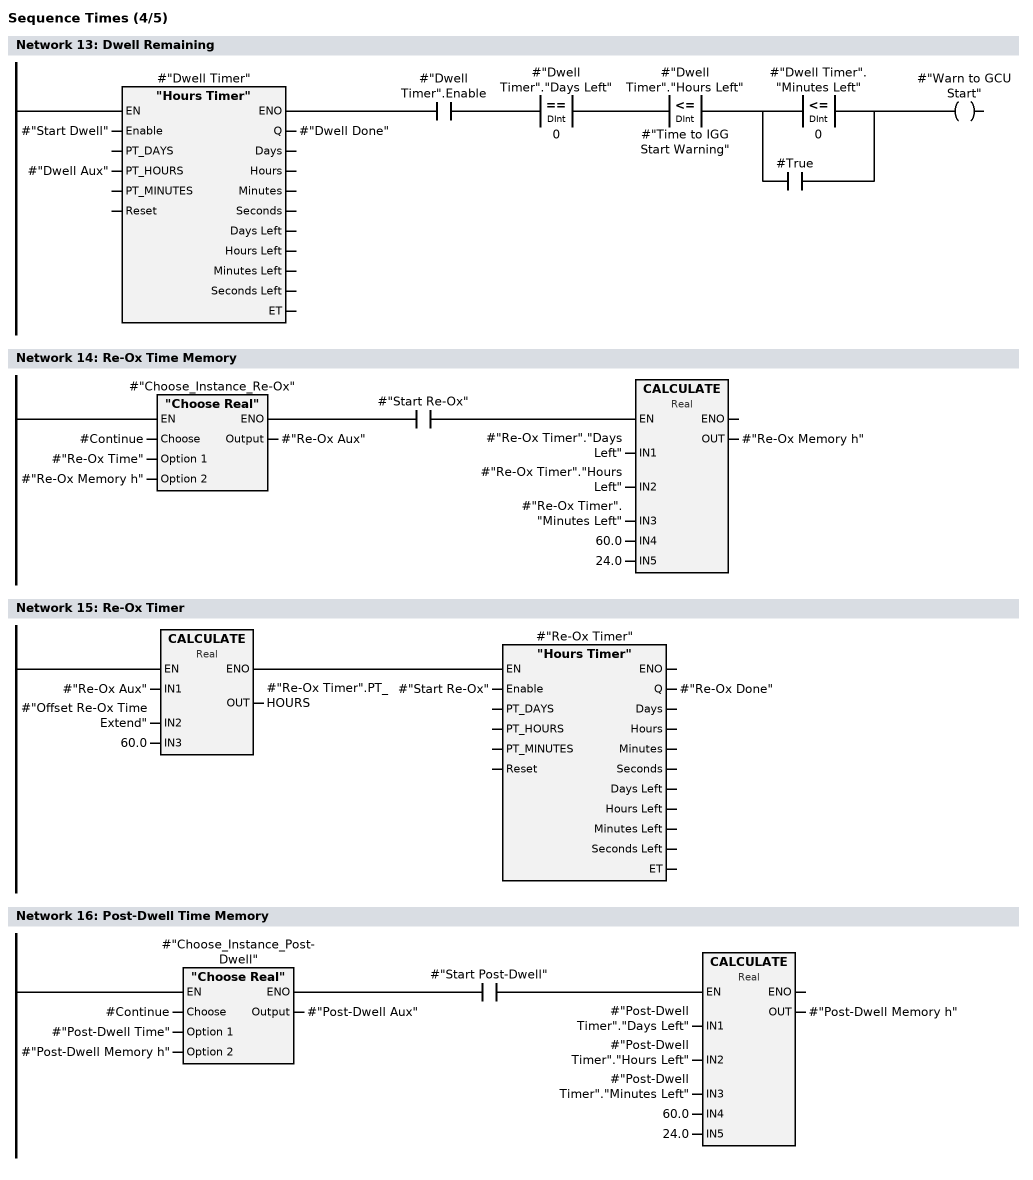
   RUNG wire#powerrail
      #"Dwell Timer"(Enable := #"Start Dwell", PT_DAYS :=, PT_HOURS := #"Dwell Aux", PT_MINUTES :=, Reset :=, Q => #"Dwell Done", Days =>, Hours =>, Minutes =>, Seconds =>, "Days Left" =>, "Hours Left" =>, "Minutes Left" =>, "Seconds Left" =>, ET =>)
      Contact( #"Dwell Timer".Enable )
      { S7_Templates := "SrcType := DInt" } EQ_Contact(in1 := #"Dwell Timer"."Days Left", in2 := 0)
      { S7_Templates := "SrcType := DInt" } LE_Contact(in1 := #"Dwell Timer"."Hours Left", in2 := #"Time to IGG Start Warning")
      wire#w1
      { S7_Templates := "SrcType := DInt" } LE_Contact(in1 := #"Dwell Timer"."Minutes Left", in2 := 0)
      wire#w2
      Coil( #"Warn to GCU Start" )
   END_RUNG
   RUNG wire#w1
      Contact( #True )
   END_RUNG wire#w2
   // the same network as SCL:
   #"Dwell Timer"(Enable := #"Start Dwell", PT_HOURS := #"Dwell Aux", Q => #"Dwell Done", ENO => #_w1);   // "Hours Timer"
   #"Warn to GCU Start" := #_w1 AND #"Dwell Timer".Enable AND (#"Dwell Timer"."Days Left" = 0) AND (#"Dwell Timer"."Hours Left" <= #"Time to IGG Start Warning") AND ((#"Dwell Timer"."Minutes Left" <= 0) OR #True);
END_REGION

REGION Network 14: Re-Ox Time Memory
   RUNG wire#powerrail
      #"Choose_Instance_Re-Ox"(Choose := #Continue, "Option 1" := #"Re-Ox Time", "Option 2" := #"Re-Ox Memory h", Output => #"Re-Ox Aux")
      Contact( #"Start Re-Ox" )
      { S7_Templates := "SrcType := Real"; S7_Expression := "(IN1*IN5)+IN2+(IN3/IN4)" } Calculate(in1 := #"Re-Ox Timer"."Days Left", in2 := #"Re-Ox Timer"."Hours Left", in3 := #"Re-Ox Timer"."Minutes Left", in4 := 60.0, in5 := 24.0, out => #"Re-Ox Memory h")
   END_RUNG
   // the same network as SCL:
   #"Choose_Instance_Re-Ox"(Choose := #Continue,   // "Choose Real"
                           "Option 1" := #"Re-Ox Time",
                           "Option 2" := #"Re-Ox Memory h",
                           Output => #"Re-Ox Aux",
                           ENO => #_w1);
   IF #_w1 AND #"Start Re-Ox" THEN
       #"Re-Ox Memory h" := (#"Re-Ox Timer"."Days Left"*24.0)+#"Re-Ox Timer"."Hours Left"+(#"Re-Ox Timer"."Minutes Left"/60.0);
   END_IF;
END_REGION

REGION Network 15: Re-Ox Timer
   RUNG wire#powerrail
      { S7_Templates := "SrcType := Real"; S7_Expression := "IN1+IN2" } Calculate(in1 := #"Re-Ox Aux", in2 := #"Offset Re-Ox Time Extend", in3 := 60.0, out => #"Re-Ox Timer".PT_HOURS)
      #"Re-Ox Timer"(Enable := #"Start Re-Ox", PT_DAYS :=, PT_HOURS :=, PT_MINUTES :=, Reset :=, Q => #"Re-Ox Done", Days =>, Hours =>, Minutes =>, Seconds =>, "Days Left" =>, "Hours Left" =>, "Minutes Left" =>, "Seconds Left" =>, ET =>)
   END_RUNG
   // the same network as SCL:
   #"Re-Ox Timer".PT_HOURS := #"Re-Ox Aux"+#"Offset Re-Ox Time Extend";
   #"Re-Ox Timer"(Enable := #"Start Re-Ox", Q => #"Re-Ox Done");   // "Hours Timer"
END_REGION

REGION Network 16: Post-Dwell Time Memory
   RUNG wire#powerrail
      #"Choose_Instance_Post-Dwell"(Choose := #Continue, "Option 1" := #"Post-Dwell Time", "Option 2" := #"Post-Dwell Memory h", Output => #"Post-Dwell Aux")
      Contact( #"Start Post-Dwell" )
      { S7_Templates := "SrcType := Real"; S7_Expression := "(IN1*IN5)+IN2+(IN3/IN4)" } Calculate(in1 := #"Post-Dwell Timer"."Days Left", in2 := #"Post-Dwell Timer"."Hours Left", in3 := #"Post-Dwell Timer"."Minutes Left", in4 := 60.0, in5 := 24.0, out => #"Post-Dwell Memory h")
   END_RUNG
   // the same network as SCL:
   #"Choose_Instance_Post-Dwell"(Choose := #Continue,   // "Choose Real"
                           "Option 1" := #"Post-Dwell Time",
                           "Option 2" := #"Post-Dwell Memory h",
                           Output => #"Post-Dwell Aux",
                           ENO => #_w1);
   IF #_w1 AND #"Start Post-Dwell" THEN
       #"Post-Dwell Memory h" := (#"Post-Dwell Timer"."Days Left"*24.0)+#"Post-Dwell Timer"."Hours Left"+(#"Post-Dwell Timer"."Minutes Left"/60.0);
   END_IF;
END_REGION

REGION Network 17: Post-Dwell Remaining
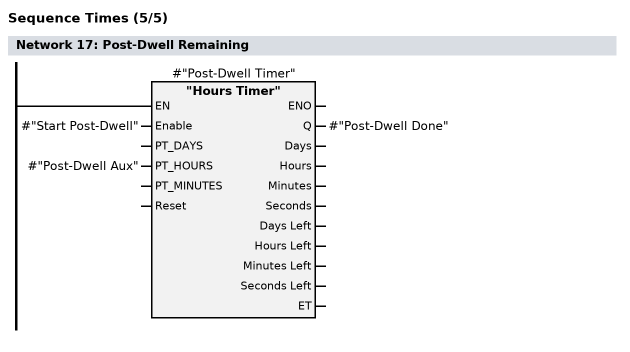
   RUNG wire#powerrail
      #"Post-Dwell Timer"(Enable := #"Start Post-Dwell", PT_DAYS :=, PT_HOURS := #"Post-Dwell Aux", PT_MINUTES :=, Reset :=, Q => #"Post-Dwell Done", Days =>, Hours =>, Minutes =>, Seconds =>, "Days Left" =>, "Hours Left" =>, "Minutes Left" =>, "Seconds Left" =>, ET =>)
   END_RUNG
   // the same network as SCL:
   #"Post-Dwell Timer"(Enable := #"Start Post-Dwell", PT_HOURS := #"Post-Dwell Aux", Q => #"Post-Dwell Done");   // "Hours Timer"
END_REGION
END_FUNCTION_BLOCK

FUNCTION_BLOCK "Days Timer"   // FB513, LAD
{ S7_Optimized_Access := 'TRUE' }
VERSION : 0.1
   VAR_INPUT
      Enable : Bool;
      PT_DAYS : Real;
   END_VAR
   VAR_OUTPUT
      Q : Bool;
      Days : Int;
      Hours : Int;
      Minutes : Int;
      Seconds : Int;
      "Days Left" : Int;
      "Hours Left" : Int;
      "Minutes Left" : Int;
      "Seconds Left" : Int;
      ET : Time;
   END_VAR
   VAR
      "Days Number" : Int;
      "Days Number_Aux" : Real;
      "Hours Number" : Int;
      "Hours Number_Aux" : Real;
      "Minutes Number" : Int;
      "Minutes Number_Aux" : Real;
      "Seconds Number" : Int;
      "Seconds Number Aux" : Real;
      "One Minute Timer" : TON_TIME;
      "One Second Timer" : TON_TIME;
      "One Second Puls" : Bool;
      "One Second Puls_aux" : Bool;
      True : Bool;
      False : Bool;
      "Enable Puls" : Bool;
   END_VAR
   VAR_TEMP   // added for the SCL form of the ladder/FBD networks
      _w1 : Bool;
      _w2 : Bool;
   END_VAR
BEGIN

REGION Network 1: True/False
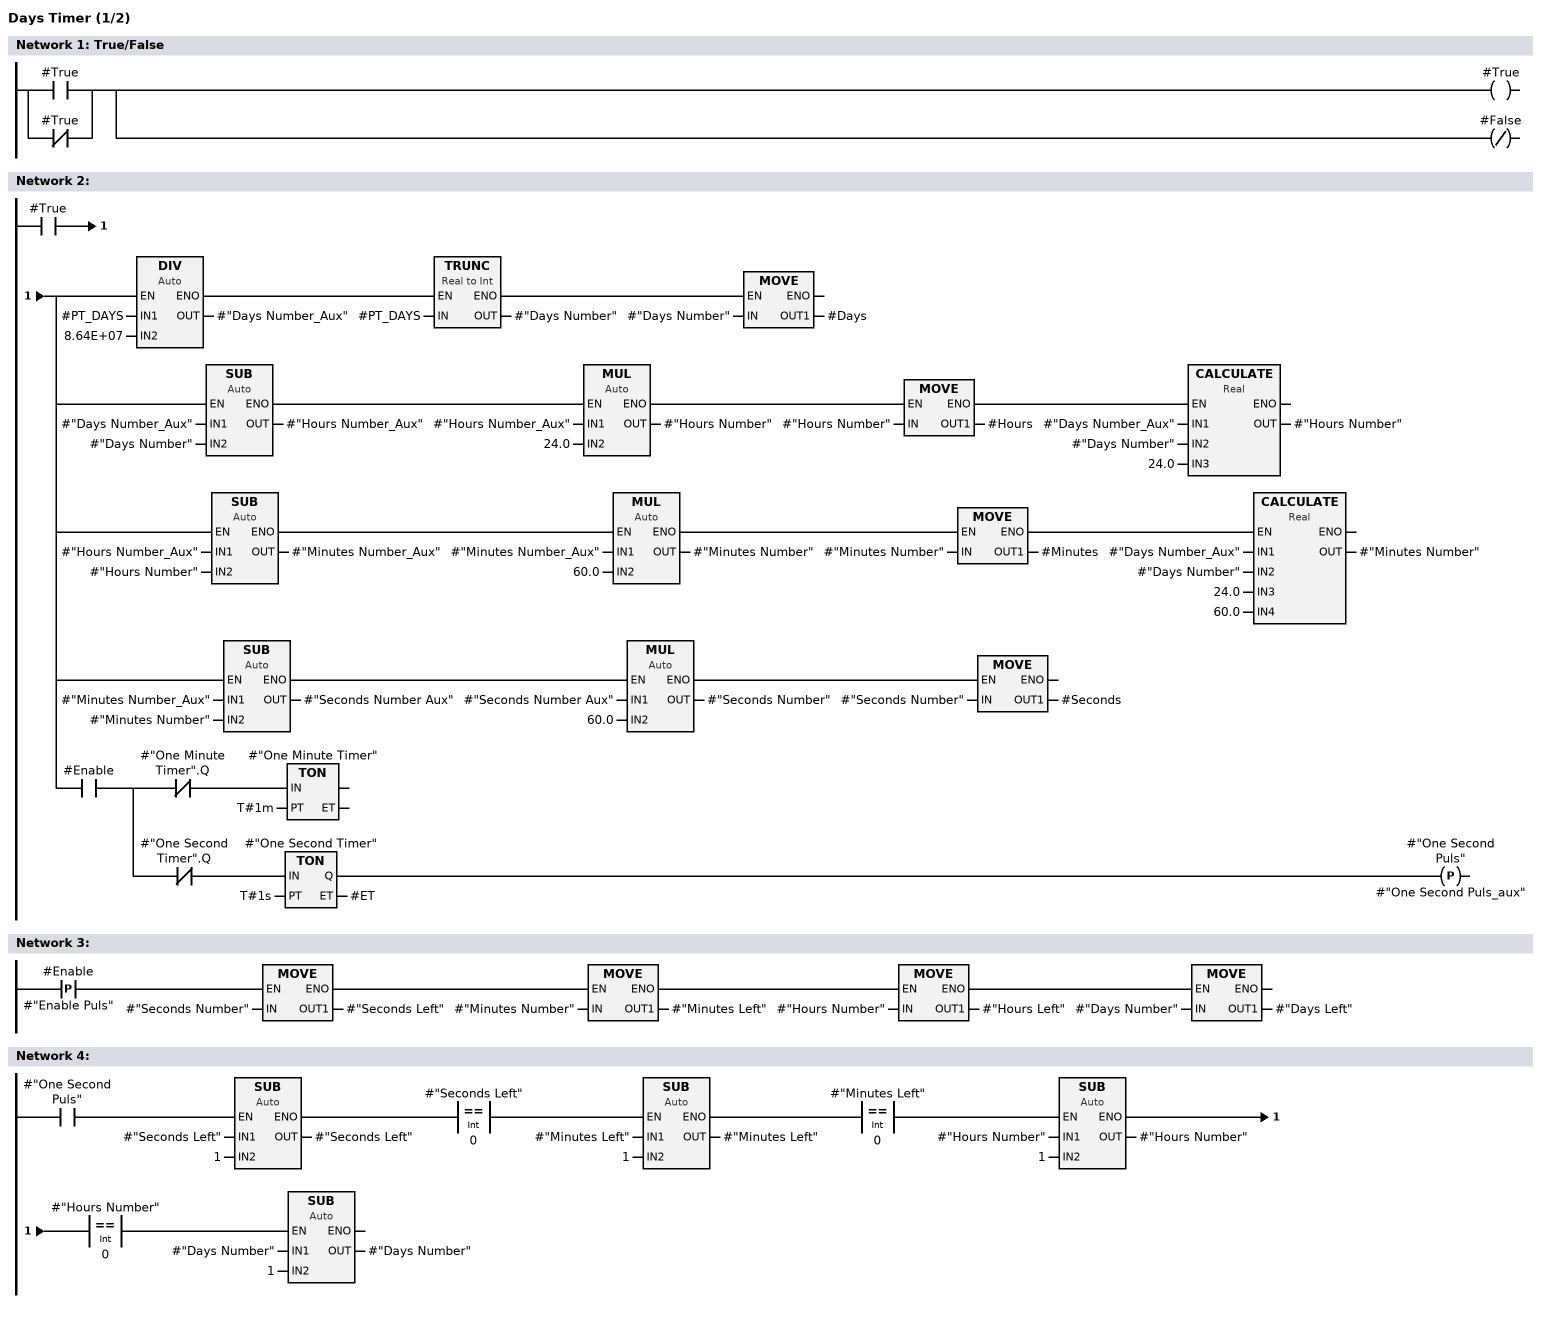
   RUNG wire#powerrail
      Contact( #True )
      wire#w1
      Coil( #True )
   END_RUNG
   RUNG wire#powerrail
      I_Contact( #True )
   END_RUNG wire#w1
   RUNG wire#w1
      I_Coil( #False )
   END_RUNG
   // the same network as SCL:
   #True := #True OR NOT #True;
   #False := NOT #True;
END_REGION

REGION Network 2
   IF #True THEN
       #"Days Number_Aux" := #PT_DAYS / 8.64E+07;
       #"Days Number" := TRUNC(#PT_DAYS);
       #Days := #"Days Number";
       #"Hours Number_Aux" := #"Days Number_Aux" - #"Days Number";
       #"Hours Number" := #"Hours Number_Aux" * 24.0;
       #Hours := #"Hours Number";
       #"Hours Number" := TRUNC((#"Days Number_Aux"-#"Days Number")*24.0);
       #"Minutes Number_Aux" := #"Hours Number_Aux" - #"Hours Number";
       #"Minutes Number" := #"Minutes Number_Aux" * 60.0;
       #Minutes := #"Minutes Number";
       #"Minutes Number" := ((#"Days Number_Aux"-(TRUNC(#"Days Number_Aux"-#"Days Number"))*24.0)-(TRUNC(#"Days Number_Aux"-(TRUNC(#"Days Number_Aux"-#"Days Number"))*24.0)))*60.0;
       #"Seconds Number Aux" := #"Minutes Number_Aux" - #"Minutes Number";
       #"Seconds Number" := #"Seconds Number Aux" * 60.0;
       #Seconds := #"Seconds Number";
   END_IF;
   #_w1 := #True AND #Enable;
   #"One Minute Timer"(IN := #_w1 AND NOT #"One Minute Timer".Q, PT := T#1m);   // TON
   #"One Second Timer"(IN := #_w1 AND NOT #"One Second Timer".Q, PT := T#1s, ET => #ET);   // TON
   #"One Second Puls" := #"One Second Timer".Q AND NOT #"One Second Puls_aux";   // rising edge
   #"One Second Puls_aux" := #"One Second Timer".Q;
END_REGION

REGION Network 3
   RUNG wire#powerrail
      P_Contact(operand := #Enable, bit := #"Enable Puls")
      Move(in := #"Seconds Number", out1 => #"Seconds Left")
      Move(in := #"Minutes Number", out1 => #"Minutes Left")
      Move(in := #"Hours Number", out1 => #"Hours Left")
      Move(in := #"Days Number", out1 => #"Days Left")
   END_RUNG
   // the same network as SCL:
   #_w1 := #Enable AND NOT #"Enable Puls";   // rising edge of #Enable
   #"Enable Puls" := #Enable;
   IF #_w1 THEN
       #"Seconds Left" := #"Seconds Number";
       #"Minutes Left" := #"Minutes Number";
       #"Hours Left" := #"Hours Number";
       #"Days Left" := #"Days Number";
   END_IF;
END_REGION

REGION Network 4
   RUNG wire#powerrail
      Contact( #"One Second Puls" )
      Sub(in1 := #"Seconds Left", in2 := 1, out => #"Seconds Left")
      { S7_Templates := "SrcType := Int" } EQ_Contact(in1 := #"Seconds Left", in2 := 0)
      Sub(in1 := #"Minutes Left", in2 := 1, out => #"Minutes Left")
      { S7_Templates := "SrcType := Int" } EQ_Contact(in1 := #"Minutes Left", in2 := 0)
      Sub(in1 := #"Hours Number", in2 := 1, out => #"Hours Number")
      { S7_Templates := "SrcType := Int" } EQ_Contact(in1 := #"Hours Number", in2 := 0)
      Sub(in1 := #"Days Number", in2 := 1, out => #"Days Number")
   END_RUNG
   // the same network as SCL:
   IF #"One Second Puls" THEN #"Seconds Left" := #"Seconds Left" - 1; END_IF;
   #_w1 := #"One Second Puls" AND (#"Seconds Left" = 0);
   IF #_w1 THEN #"Minutes Left" := #"Minutes Left" - 1; END_IF;
   #_w2 := #_w1 AND (#"Minutes Left" = 0);
   IF #_w2 THEN #"Hours Number" := #"Hours Number" - 1; END_IF;
   IF #_w2 AND (#"Hours Number" = 0) THEN #"Days Number" := #"Days Number" - 1; END_IF;
END_REGION

REGION Network 5
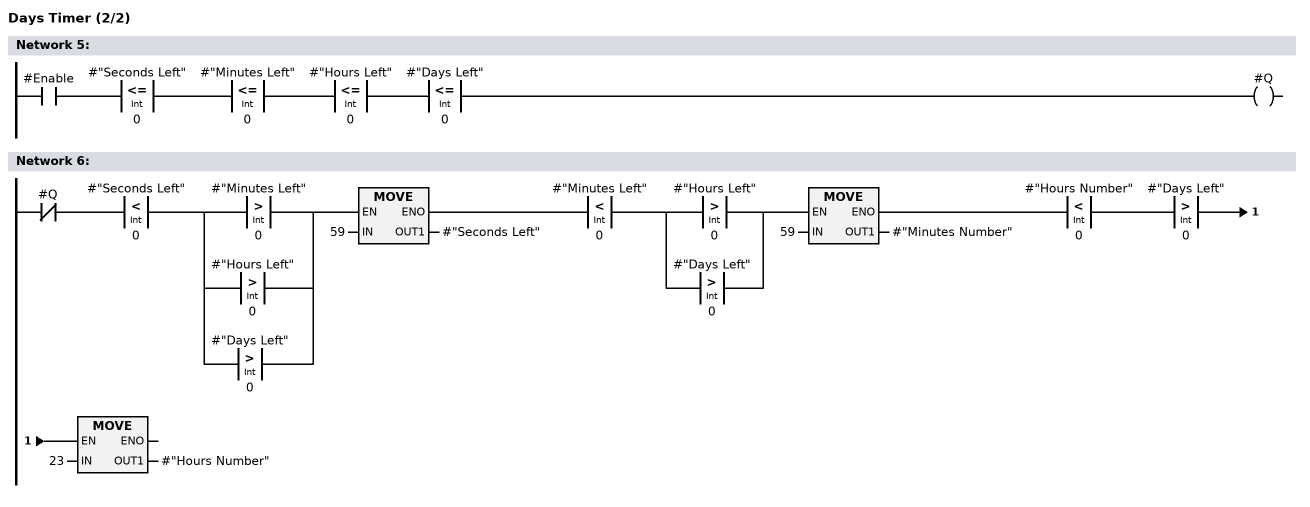
   RUNG wire#powerrail
      Contact( #Enable )
      { S7_Templates := "SrcType := Int" } LE_Contact(in1 := #"Seconds Left", in2 := 0)
      { S7_Templates := "SrcType := Int" } LE_Contact(in1 := #"Minutes Left", in2 := 0)
      { S7_Templates := "SrcType := Int" } LE_Contact(in1 := #"Hours Left", in2 := 0)
      { S7_Templates := "SrcType := Int" } LE_Contact(in1 := #"Days Left", in2 := 0)
      Coil( #Q )
   END_RUNG
   // the same network as SCL:
   #Q := #Enable AND (#"Seconds Left" <= 0) AND (#"Minutes Left" <= 0) AND (#"Hours Left" <= 0) AND (#"Days Left" <= 0);
END_REGION

REGION Network 6
   RUNG wire#powerrail
      I_Contact( #Q )
      { S7_Templates := "SrcType := Int" } LT_Contact(in1 := #"Seconds Left", in2 := 0)
      wire#w1
      { S7_Templates := "SrcType := Int" } GT_Contact(in1 := #"Minutes Left", in2 := 0)
      wire#w2
      Move(in := 59, out1 => #"Seconds Left")
      { S7_Templates := "SrcType := Int" } LT_Contact(in1 := #"Minutes Left", in2 := 0)
      wire#w3
      { S7_Templates := "SrcType := Int" } GT_Contact(in1 := #"Hours Left", in2 := 0)
      wire#w4
      Move(in := 59, out1 => #"Minutes Number")
      { S7_Templates := "SrcType := Int" } LT_Contact(in1 := #"Hours Number", in2 := 0)
      { S7_Templates := "SrcType := Int" } GT_Contact(in1 := #"Days Left", in2 := 0)
      Move(in := 23, out1 => #"Hours Number")
   END_RUNG
   RUNG wire#w1
      { S7_Templates := "SrcType := Int" } GT_Contact(in1 := #"Hours Left", in2 := 0)
   END_RUNG wire#w2
   RUNG wire#w1
      { S7_Templates := "SrcType := Int" } GT_Contact(in1 := #"Days Left", in2 := 0)
   END_RUNG wire#w2
   RUNG wire#w3
      { S7_Templates := "SrcType := Int" } GT_Contact(in1 := #"Days Left", in2 := 0)
   END_RUNG wire#w4
   // the same network as SCL:
   #_w1 := NOT #Q AND (#"Seconds Left" < 0) AND ((#"Minutes Left" > 0) OR (#"Hours Left" > 0) OR (#"Days Left" > 0));
   IF #_w1 THEN #"Seconds Left" := 59; END_IF;
   #_w2 := #_w1 AND (#"Minutes Left" < 0) AND ((#"Hours Left" > 0) OR (#"Days Left" > 0));
   IF #_w2 THEN #"Minutes Number" := 59; END_IF;
   IF #_w2 AND (#"Hours Number" < 0) AND (#"Days Left" > 0) THEN #"Hours Number" := 23; END_IF;
END_REGION
END_FUNCTION_BLOCK

FUNCTION_BLOCK "Hours Timer"   // FB514, LAD
{ S7_Optimized_Access := 'TRUE' }
VERSION : 0.1
   VAR_INPUT
      Enable : Bool;
      PT_DAYS : Real;
      PT_HOURS : Real;
      PT_MINUTES : Real;
      Reset : Bool;
   END_VAR
   VAR_OUTPUT
      Q : Bool;
      Days : DInt;
      Hours : DInt;
      Minutes : DInt;
      Seconds : DInt;
      "Days Left" : DInt;
      "Hours Left" : DInt;
      "Minutes Left" : DInt;
      "Seconds Left" : DInt;
      ET : Time;
   END_VAR
   VAR
      "Days Number" : Int;
      "Days Number_Aux" : Real;
      "Hours Number" : Int;
      "Hours Number_Real" : Real;
      "Hours Number_Aux" : Real;
      "Minutes Number" : Int;
      "Minutes Number_Real" : Real;
      "Minutes Number_Aux" : Real;
      "Seconds Number" : Int;
      "Seconds Number Real" : Real;
      "Seconds Number Aux" : Real;
      "One Minute Timer" : TON_TIME;
      "One Second Timer" : TON_TIME;
      "One Second Puls" : Bool;
      "One Second Puls_aux" : Bool;
      True : Bool;
      False : Bool;
      "Enable Puls" : Bool;
      "Enable Puls N" : Bool;
      "One Second Puls TP" : TP_TIME;
   END_VAR
   VAR_TEMP   // added for the SCL form of the ladder/FBD networks
      _w1 : Bool;
      _w2 : Bool;
      _w3 : Bool;
      _w4 : Bool;
   END_VAR
BEGIN

REGION Network 1: True/False
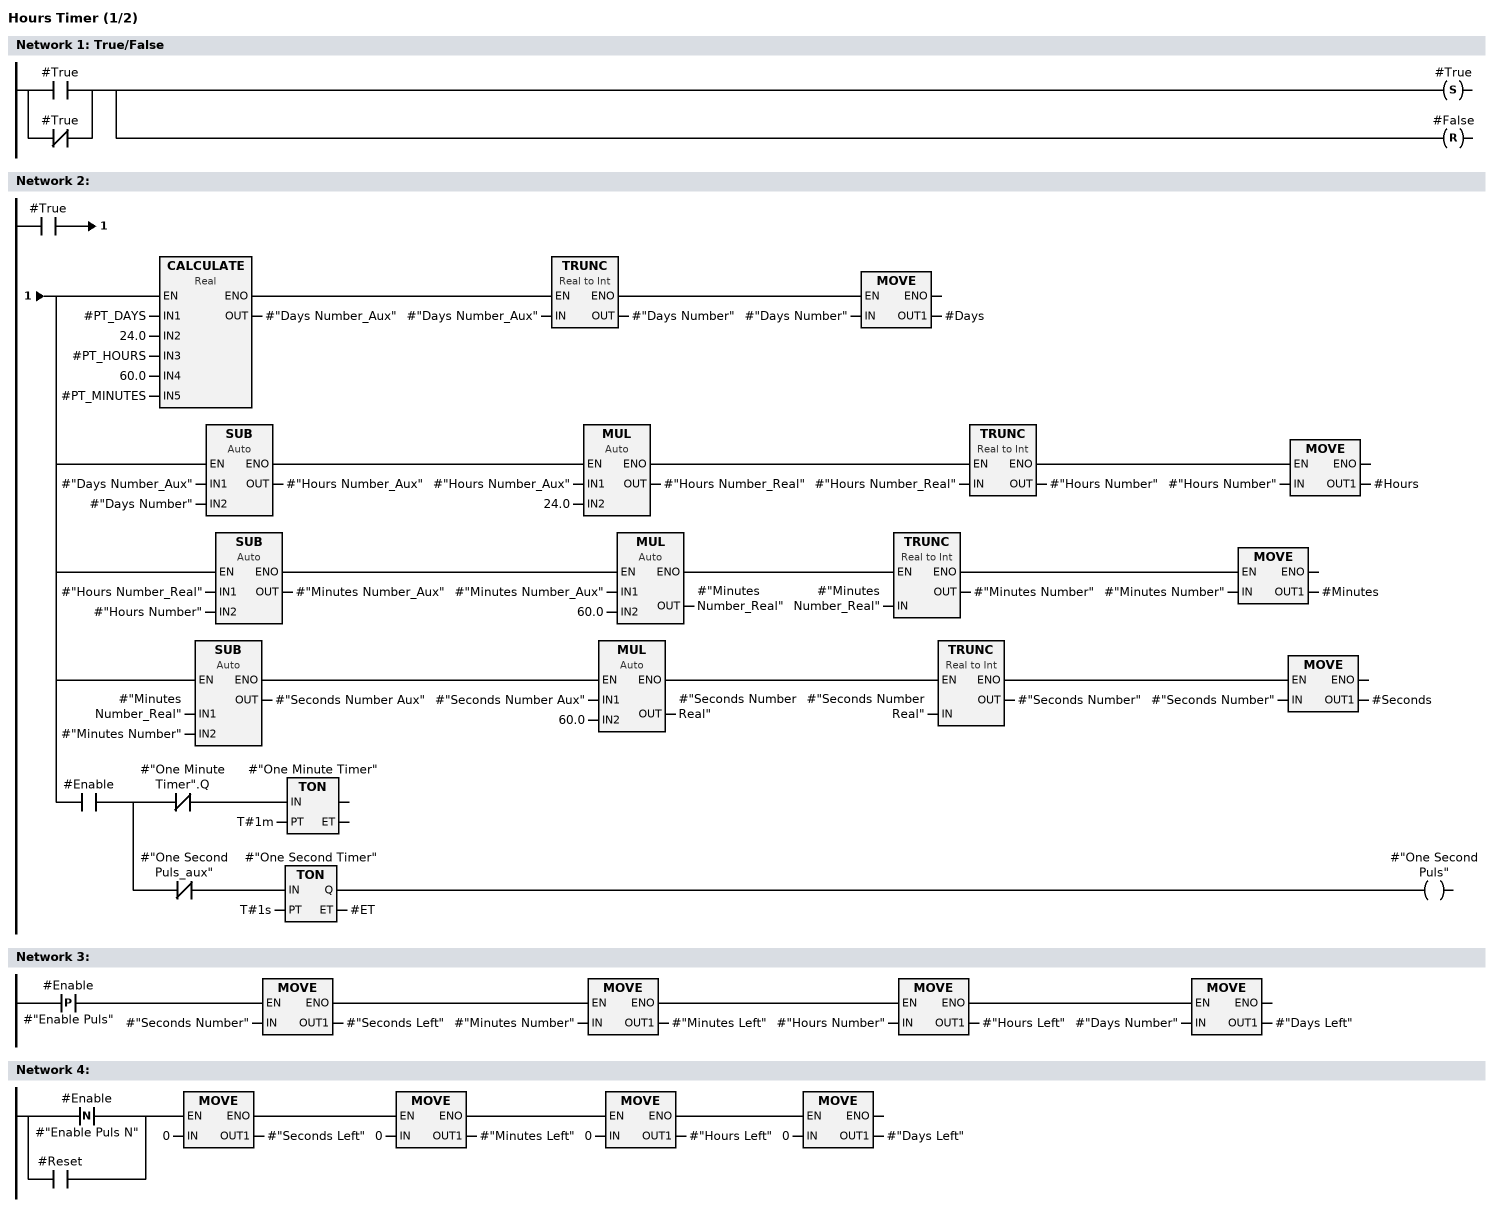
   RUNG wire#powerrail
      Contact( #True )
      wire#w1
      S_Coil( #True )
   END_RUNG
   RUNG wire#powerrail
      I_Contact( #True )
   END_RUNG wire#w1
   RUNG wire#w1
      R_Coil( #False )
   END_RUNG
   // the same network as SCL:
   #_w1 := #True OR NOT #True;
   IF #_w1 THEN
       #True := TRUE;
       #False := FALSE;
   END_IF;
END_REGION

REGION Network 2
   IF #True THEN
       #"Days Number_Aux" := #PT_DAYS+(#PT_HOURS/24.0)+(#PT_MINUTES/60.0);
       #"Days Number" := TRUNC(#"Days Number_Aux");
       #Days := #"Days Number";
       #"Hours Number_Aux" := #"Days Number_Aux" - #"Days Number";
       #"Hours Number_Real" := #"Hours Number_Aux" * 24.0;
       #"Hours Number" := TRUNC(#"Hours Number_Real");
       #Hours := #"Hours Number";
       #"Minutes Number_Aux" := #"Hours Number_Real" - #"Hours Number";
       #"Minutes Number_Real" := #"Minutes Number_Aux" * 60.0;
       #"Minutes Number" := TRUNC(#"Minutes Number_Real");
       #Minutes := #"Minutes Number";
       #"Seconds Number Aux" := #"Minutes Number_Real" - #"Minutes Number";
       #"Seconds Number Real" := #"Seconds Number Aux" * 60.0;
       #"Seconds Number" := TRUNC(#"Seconds Number Real");
       #Seconds := #"Seconds Number";
   END_IF;
   #_w1 := #True AND #Enable;
   #"One Minute Timer"(IN := #_w1 AND NOT #"One Minute Timer".Q, PT := T#1m);   // TON
   #"One Second Timer"(IN := #_w1 AND NOT #"One Second Puls_aux", PT := T#1s, ET => #ET);   // TON
   #"One Second Puls" := #"One Second Timer".Q;
END_REGION

REGION Network 3
   RUNG wire#powerrail
      P_Contact(operand := #Enable, bit := #"Enable Puls")
      Move(in := #"Seconds Number", out1 => #"Seconds Left")
      Move(in := #"Minutes Number", out1 => #"Minutes Left")
      Move(in := #"Hours Number", out1 => #"Hours Left")
      Move(in := #"Days Number", out1 => #"Days Left")
   END_RUNG
   // the same network as SCL:
   #_w1 := #Enable AND NOT #"Enable Puls";   // rising edge of #Enable
   #"Enable Puls" := #Enable;
   IF #_w1 THEN
       #"Seconds Left" := #"Seconds Number";
       #"Minutes Left" := #"Minutes Number";
       #"Hours Left" := #"Hours Number";
       #"Days Left" := #"Days Number";
   END_IF;
END_REGION

REGION Network 4
   RUNG wire#powerrail
      N_Contact(operand := #Enable, bit := #"Enable Puls N")
      wire#w1
      Move(in := 0, out1 => #"Seconds Left")
      Move(in := 0, out1 => #"Minutes Left")
      Move(in := 0, out1 => #"Hours Left")
      Move(in := 0, out1 => #"Days Left")
   END_RUNG
   RUNG wire#powerrail
      Contact( #Reset )
   END_RUNG wire#w1
   // the same network as SCL:
   #_w1 := NOT #Enable AND #"Enable Puls N";   // falling edge of #Enable
   #"Enable Puls N" := #Enable;
   IF #_w1 OR #Reset THEN
       #"Seconds Left" := 0;
       #"Minutes Left" := 0;
       #"Hours Left" := 0;
       #"Days Left" := 0;
   END_IF;
END_REGION

REGION Network 5: Cout Down
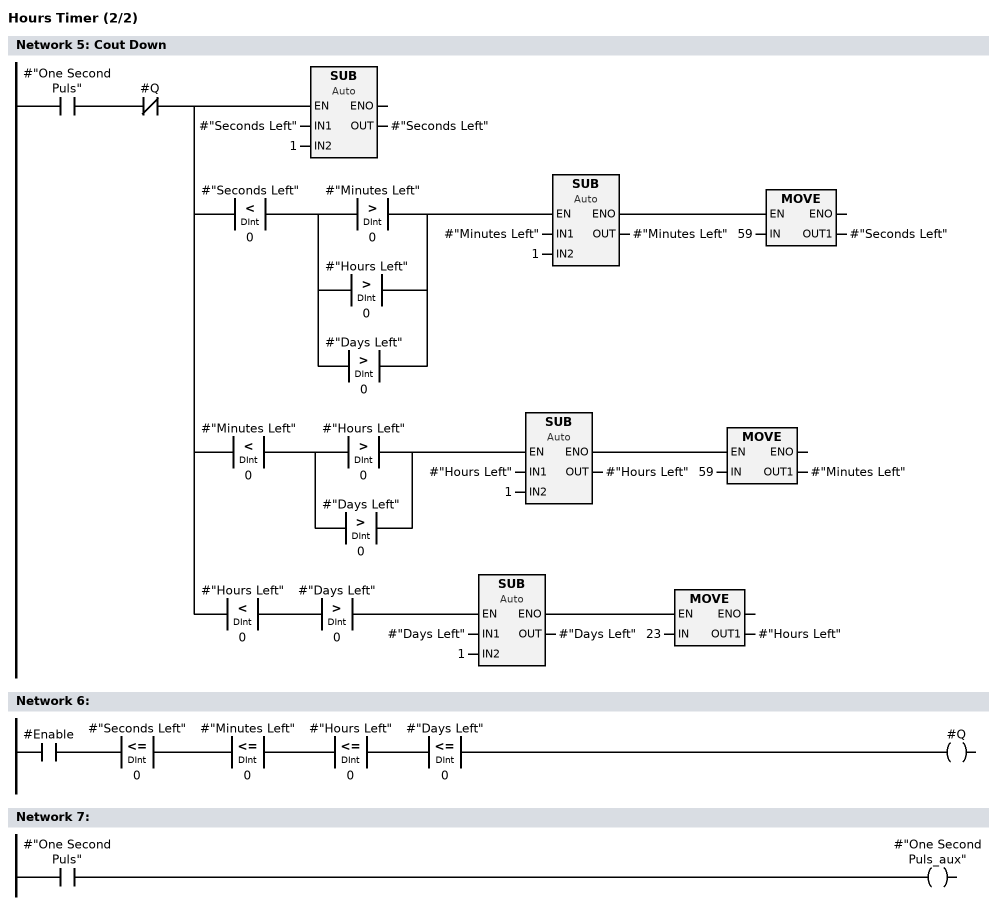
   RUNG wire#powerrail
      Contact( #"One Second Puls" )
      I_Contact( #Q )
      wire#w1
      Sub(in1 := #"Seconds Left", in2 := 1, out => #"Seconds Left")
   END_RUNG
   RUNG wire#w1
      { S7_Templates := "SrcType := DInt" } LT_Contact(in1 := #"Seconds Left", in2 := 0)
      wire#w2
      { S7_Templates := "SrcType := DInt" } GT_Contact(in1 := #"Minutes Left", in2 := 0)
      wire#w3
      Sub(in1 := #"Minutes Left", in2 := 1, out => #"Minutes Left")
      Move(in := 59, out1 => #"Seconds Left")
   END_RUNG
   RUNG wire#w2
      { S7_Templates := "SrcType := DInt" } GT_Contact(in1 := #"Hours Left", in2 := 0)
   END_RUNG wire#w3
   RUNG wire#w2
      { S7_Templates := "SrcType := DInt" } GT_Contact(in1 := #"Days Left", in2 := 0)
   END_RUNG wire#w3
   RUNG wire#w1
      { S7_Templates := "SrcType := DInt" } LT_Contact(in1 := #"Minutes Left", in2 := 0)
      wire#w4
      { S7_Templates := "SrcType := DInt" } GT_Contact(in1 := #"Hours Left", in2 := 0)
      wire#w5
      Sub(in1 := #"Hours Left", in2 := 1, out => #"Hours Left")
      Move(in := 59, out1 => #"Minutes Left")
   END_RUNG
   RUNG wire#w4
      { S7_Templates := "SrcType := DInt" } GT_Contact(in1 := #"Days Left", in2 := 0)
   END_RUNG wire#w5
   RUNG wire#w1
      { S7_Templates := "SrcType := DInt" } LT_Contact(in1 := #"Hours Left", in2 := 0)
      { S7_Templates := "SrcType := DInt" } GT_Contact(in1 := #"Days Left", in2 := 0)
      Sub(in1 := #"Days Left", in2 := 1, out => #"Days Left")
      Move(in := 23, out1 => #"Hours Left")
   END_RUNG
   // the same network as SCL:
   #_w1 := #"One Second Puls" AND NOT #Q;
   IF #_w1 THEN #"Seconds Left" := #"Seconds Left" - 1; END_IF;
   #_w2 := #_w1 AND (#"Seconds Left" < 0) AND ((#"Minutes Left" > 0) OR (#"Hours Left" > 0) OR (#"Days Left" > 0));
   IF #_w2 THEN
       #"Minutes Left" := #"Minutes Left" - 1;
       #"Seconds Left" := 59;
   END_IF;
   #_w3 := #_w1 AND (#"Minutes Left" < 0) AND ((#"Hours Left" > 0) OR (#"Days Left" > 0));
   IF #_w3 THEN
       #"Hours Left" := #"Hours Left" - 1;
       #"Minutes Left" := 59;
   END_IF;
   #_w4 := #_w1 AND (#"Hours Left" < 0) AND (#"Days Left" > 0);
   IF #_w4 THEN
       #"Days Left" := #"Days Left" - 1;
       #"Hours Left" := 23;
   END_IF;
END_REGION

REGION Network 6
   RUNG wire#powerrail
      Contact( #Enable )
      { S7_Templates := "SrcType := DInt" } LE_Contact(in1 := #"Seconds Left", in2 := 0)
      { S7_Templates := "SrcType := DInt" } LE_Contact(in1 := #"Minutes Left", in2 := 0)
      { S7_Templates := "SrcType := DInt" } LE_Contact(in1 := #"Hours Left", in2 := 0)
      { S7_Templates := "SrcType := DInt" } LE_Contact(in1 := #"Days Left", in2 := 0)
      Coil( #Q )
   END_RUNG
   // the same network as SCL:
   #Q := #Enable AND (#"Seconds Left" <= 0) AND (#"Minutes Left" <= 0) AND (#"Hours Left" <= 0) AND (#"Days Left" <= 0);
END_REGION

REGION Network 7
   RUNG wire#powerrail
      Contact( #"One Second Puls" )
      Coil( #"One Second Puls_aux" )
   END_RUNG
   // the same network as SCL:
   #"One Second Puls_aux" := #"One Second Puls";
END_REGION
END_FUNCTION_BLOCK

FUNCTION_BLOCK "Animation"   // FB515, LAD
{ S7_Optimized_Access := 'TRUE' }
VERSION : 0.1
   VAR_INPUT
      Run : Bool;
      Revert : Bool := true;
      "States Number" : Int := 10;
      Period : Time := T#250ms;
   END_VAR
   VAR_OUTPUT
      Animation : Int;
   END_VAR
   VAR RETAIN
      "Animation State" : CTU_INT;
      Reset : Bool;
   END_VAR
   VAR
      "Revert Aux" : Bool;
      LD : Bool;
      OFF : TON_TIME;
      ON : TON_TIME;
   END_VAR
BEGIN

REGION Network 1
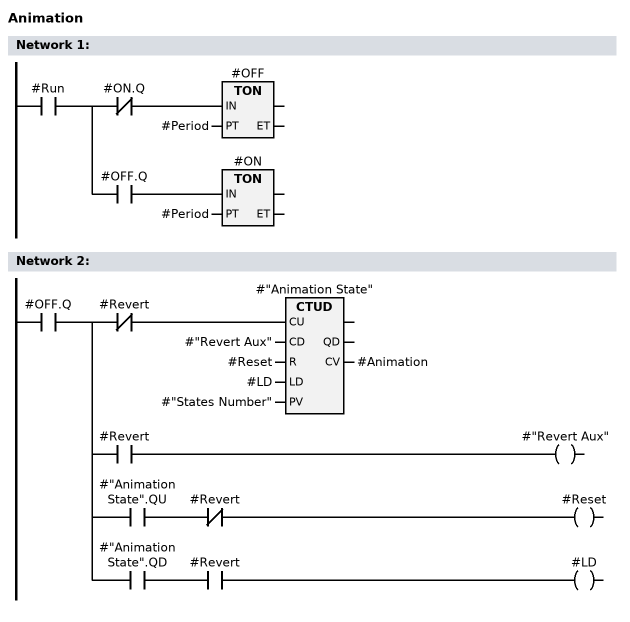
   #OFF(IN := #Run AND NOT #ON.Q, PT := #Period);   // TON
   #ON(IN := #Run AND #OFF.Q, PT := #Period);   // TON
END_REGION

REGION Network 2
   #"Animation State"(CU := #OFF.Q AND NOT #Revert,   // CTUD
                      CD := #"Revert Aux",
                      R := #Reset,
                      LD := #LD,
                      PV := #"States Number",
                      CV => #Animation);
   #"Revert Aux" := #OFF.Q AND #Revert;
   #Reset := #OFF.Q AND #"Animation State".QU AND NOT #Revert;
   #LD := #OFF.Q AND #"Animation State".QD AND #Revert;
END_REGION
END_FUNCTION_BLOCK

FUNCTION_BLOCK "DInt to Real Calcul #Out := (INT_TO_REAL((#IN1 + #IN2 + #IN3) - (#IN4 + #IN5 + #IN6)) / #IN7)"   // FB516, LAD
{ S7_Optimized_Access := 'TRUE' }